(* Logix 5000 project; controller Joltek_RA_5069PLC002 vendor 1 type 14 code 226 rev 34.15; software revision 34.04 *) (continued)
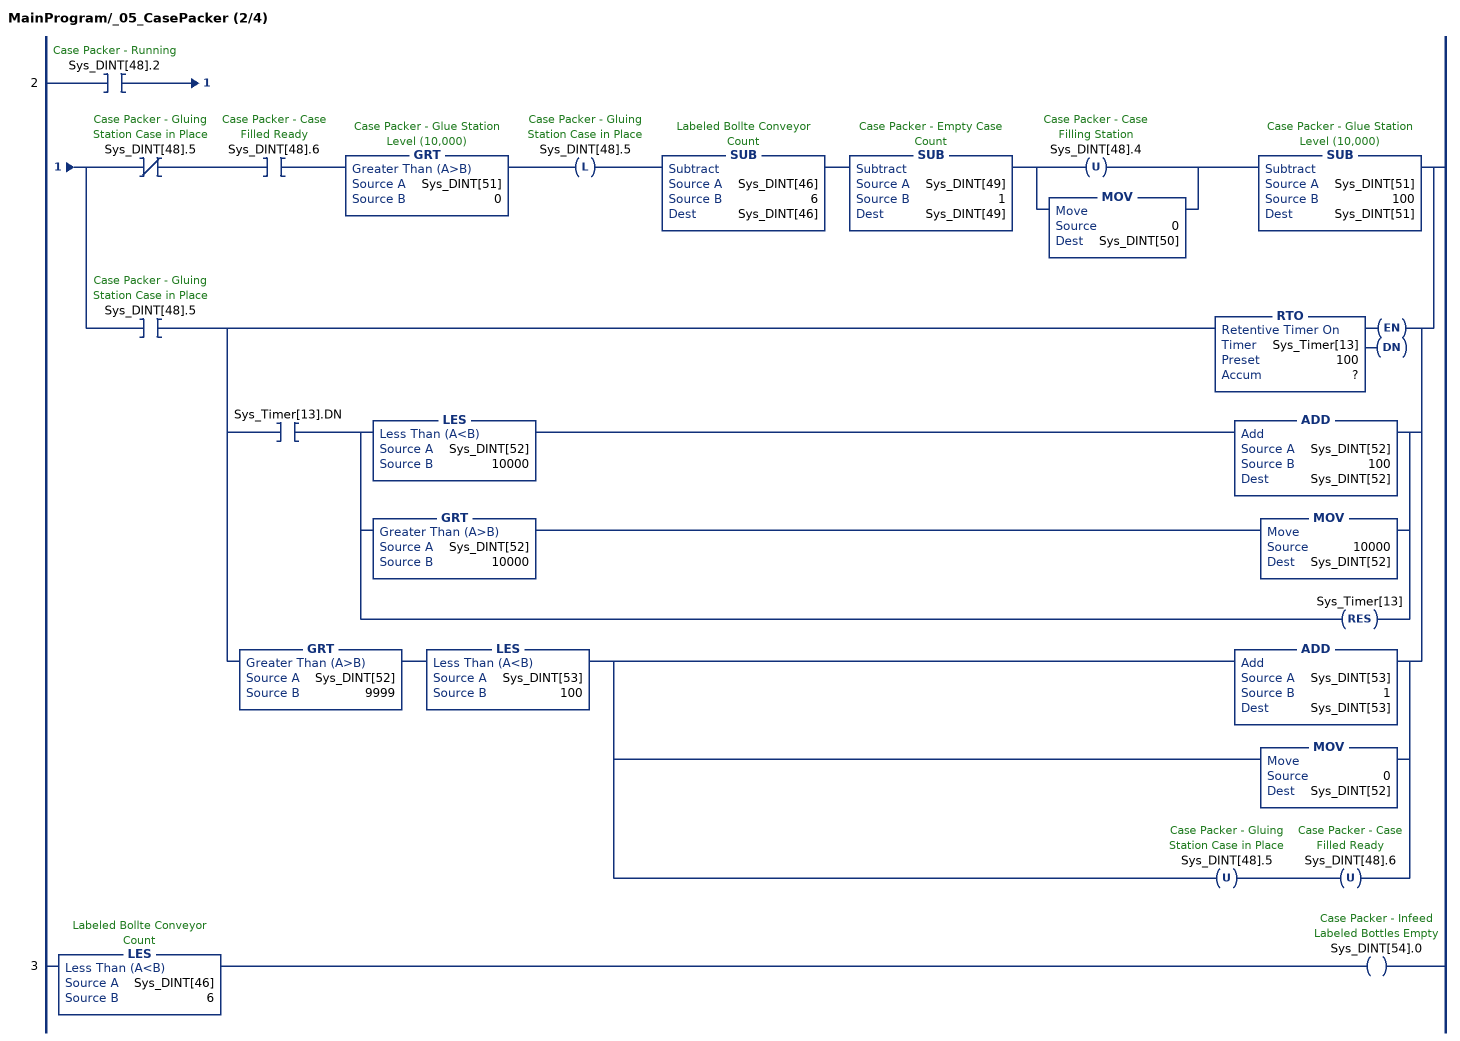
   2: XIC(Sys_DINT[48].2)[XIO(Sys_DINT[48].5) XIC(Sys_DINT[48].6) GRT(Sys_DINT[51],0) OTL(Sys_DINT[48].5) SUB(Sys_DINT[46],6,Sys_DINT[46]) SUB(Sys_DINT[49],1,Sys_DINT[49]) [OTU(Sys_DINT[48].4) ,MOV(0,Sys_DINT[50]) ] SUB(Sys_DINT[51],100,Sys_DINT[51]) ,XIC(Sys_DINT[48].5) [RTO(Sys_Timer[13],?,?) ,XIC(Sys_Timer[13].DN) [LES(Sys_DINT[52],10000) ADD(Sys_DINT[52],100,Sys_DINT[52]) ,GRT(Sys_DINT[52],10000) MOV(10000,Sys_DINT[52]) ,RES(Sys_Timer[13]) ] ,GRT(Sys_DINT[52],9999) LES(Sys_DINT[53],100) [ADD(Sys_DINT[53],1,Sys_DINT[53]) ,MOV(0,Sys_DINT[52]) ,OTU(Sys_DINT[48].5) OTU(Sys_DINT[48].6) ] ] ];
   3: LES(Sys_DINT[46],6)OTE(Sys_DINT[54].0);
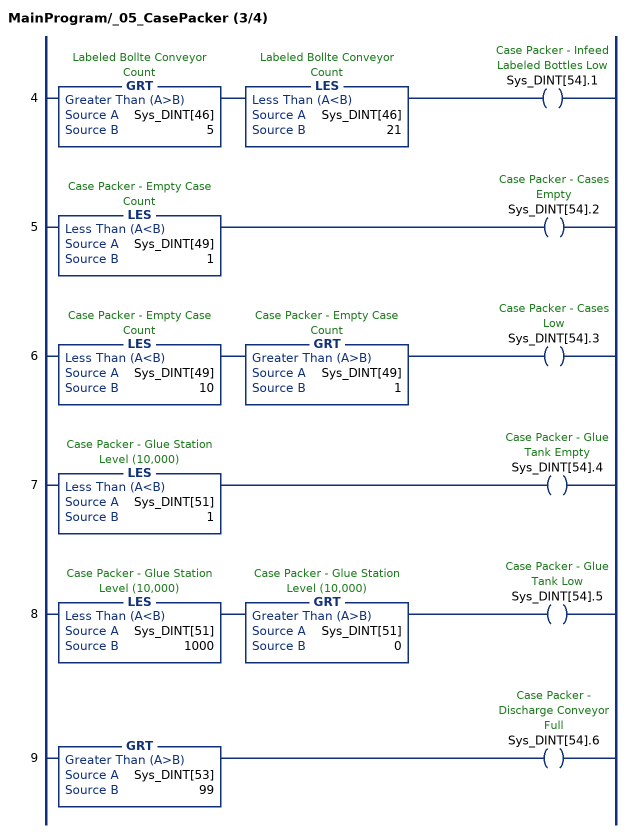
   4: GRT(Sys_DINT[46],5)LES(Sys_DINT[46],21)OTE(Sys_DINT[54].1);
   5: LES(Sys_DINT[49],1)OTE(Sys_DINT[54].2);
   6: LES(Sys_DINT[49],10)GRT(Sys_DINT[49],1)OTE(Sys_DINT[54].3);
   7: LES(Sys_DINT[51],1)OTE(Sys_DINT[54].4);
   8: LES(Sys_DINT[51],1000)GRT(Sys_DINT[51],0)OTE(Sys_DINT[54].5);
   9: GRT(Sys_DINT[53],99)OTE(Sys_DINT[54].6);
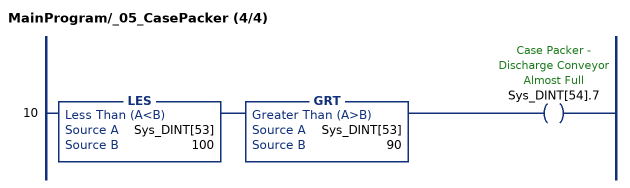
   10: LES(Sys_DINT[53],100)GRT(Sys_DINT[53],90)OTE(Sys_DINT[54].7);
END_ROUTINE

ROUTINE _06_Palletizer   (* ladder *)
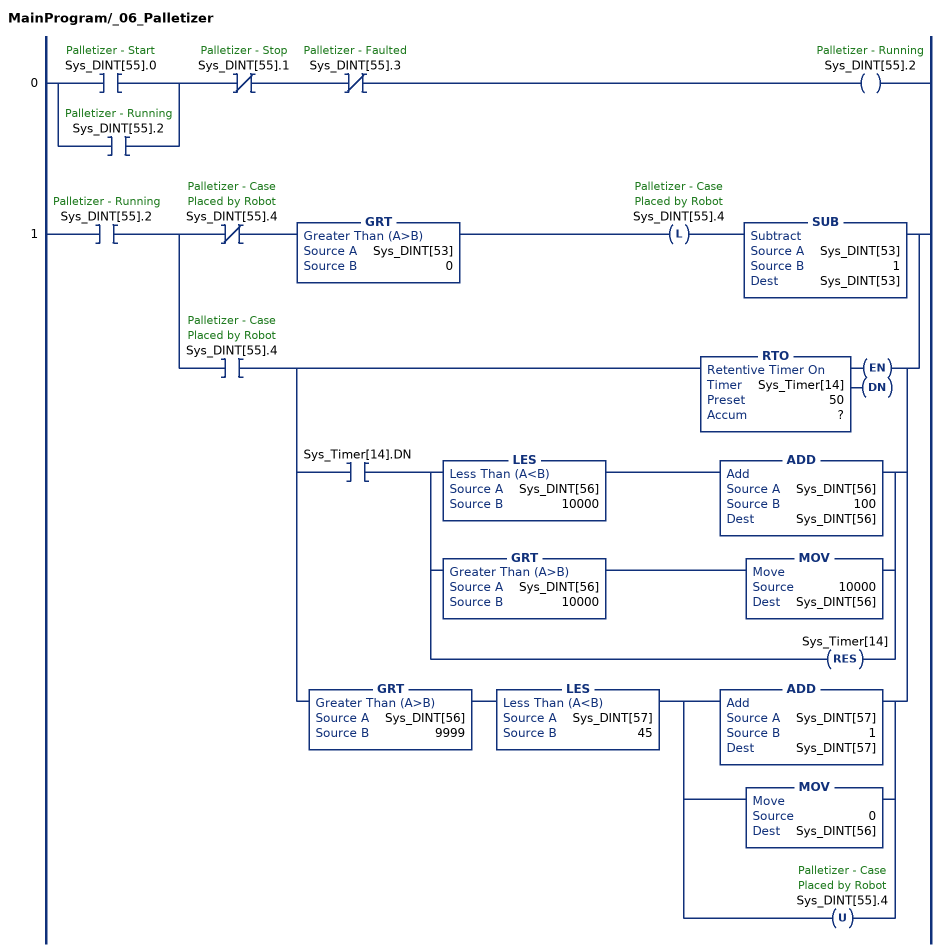
   0: [XIC(Sys_DINT[55].0) ,XIC(Sys_DINT[55].2) ]XIO(Sys_DINT[55].1)XIO(Sys_DINT[55].3)OTE(Sys_DINT[55].2);
   1: XIC(Sys_DINT[55].2)[XIO(Sys_DINT[55].4) GRT(Sys_DINT[53],0) OTL(Sys_DINT[55].4) SUB(Sys_DINT[53],1,Sys_DINT[53]) ,XIC(Sys_DINT[55].4) [RTO(Sys_Timer[14],?,?) ,XIC(Sys_Timer[14].DN) [LES(Sys_DINT[56],10000) ADD(Sys_DINT[56],100,Sys_DINT[56]) ,GRT(Sys_DINT[56],10000) MOV(10000,Sys_DINT[56]) ,RES(Sys_Timer[14]) ] ,GRT(Sys_DINT[56],9999) LES(Sys_DINT[57],45) [ADD(Sys_DINT[57],1,Sys_DINT[57]) ,MOV(0,Sys_DINT[56]) ,OTU(Sys_DINT[55].4) ] ] ];
END_ROUTINE

ROUTINE _50_HMI_Interface   (* ladder *)
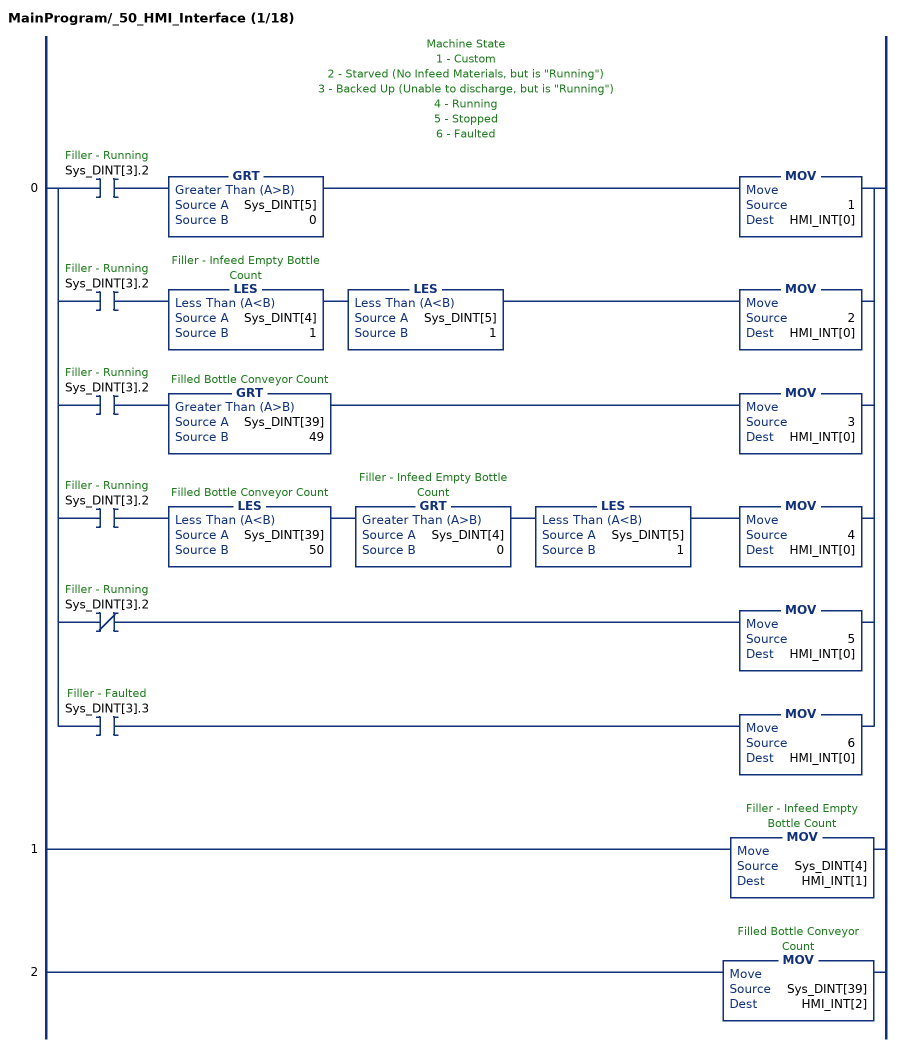
   // Machine State
   // 1 - Custom
   // 2 - Starved (No Infeed Materials, but is "Running")
   // 3 - Backed Up (Unable to discharge, but is "Running")
   // 4 - Running
   // 5 - Stopped
   // 6 - Faulted
   0: [XIC(Sys_DINT[3].2) GRT(Sys_DINT[5],0) MOV(1,HMI_INT[0]) ,XIC(Sys_DINT[3].2) LES(Sys_DINT[4],1) LES(Sys_DINT[5],1) MOV(2,HMI_INT[0]) ,XIC(Sys_DINT[3].2) GRT(Sys_DINT[39],49) MOV(3,HMI_INT[0]) ,XIC(Sys_DINT[3].2) LES(Sys_DINT[39],50) GRT(Sys_DINT[4],0) LES(Sys_DINT[5],1) MOV(4,HMI_INT[0]) ,XIO(Sys_DINT[3].2) MOV(5,HMI_INT[0]) ,XIC(Sys_DINT[3].3) MOV(6,HMI_INT[0]) ];
   1: MOV(Sys_DINT[4],HMI_INT[1]);
   2: MOV(Sys_DINT[39],HMI_INT[2]);
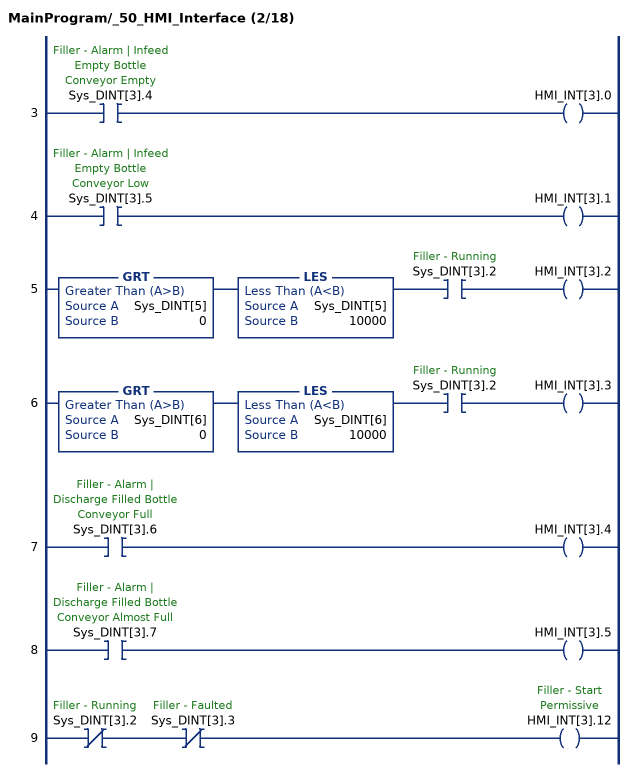
   3: XIC(Sys_DINT[3].4)OTE(HMI_INT[3].0);
   4: XIC(Sys_DINT[3].5)OTE(HMI_INT[3].1);
   5: GRT(Sys_DINT[5],0)LES(Sys_DINT[5],10000)XIC(Sys_DINT[3].2)OTE(HMI_INT[3].2);
   6: GRT(Sys_DINT[6],0)LES(Sys_DINT[6],10000)XIC(Sys_DINT[3].2)OTE(HMI_INT[3].3);
   7: XIC(Sys_DINT[3].6)OTE(HMI_INT[3].4);
   8: XIC(Sys_DINT[3].7)OTE(HMI_INT[3].5);
   9: XIO(Sys_DINT[3].2)XIO(Sys_DINT[3].3)OTE(HMI_INT[3].12);
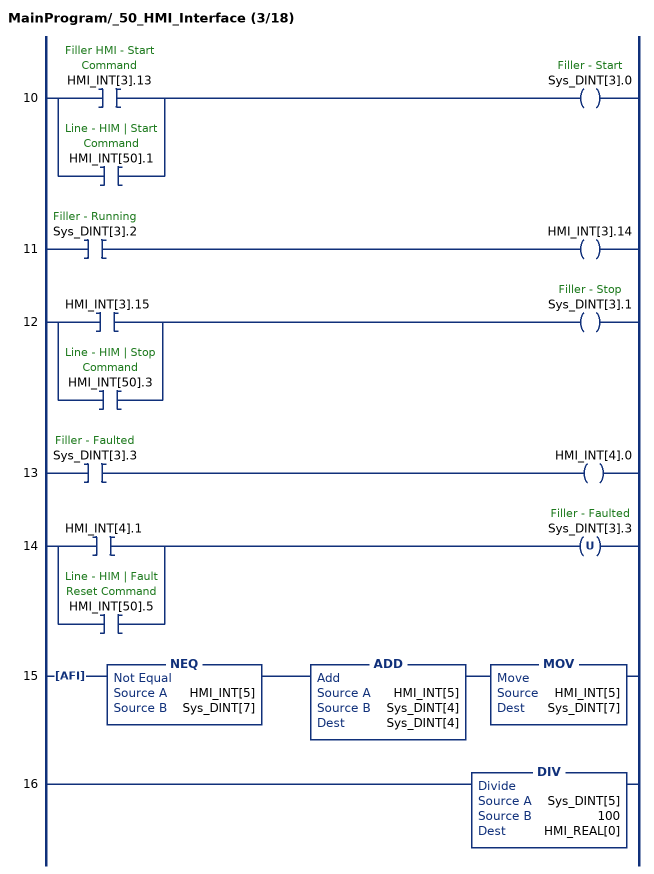
   10: [XIC(HMI_INT[3].13) ,XIC(HMI_INT[50].1) ]OTE(Sys_DINT[3].0);
   11: XIC(Sys_DINT[3].2)OTE(HMI_INT[3].14);
   12: [XIC(HMI_INT[3].15) ,XIC(HMI_INT[50].3) ]OTE(Sys_DINT[3].1);
   13: XIC(Sys_DINT[3].3)OTE(HMI_INT[4].0);
   14: [XIC(HMI_INT[4].1) ,XIC(HMI_INT[50].5) ]OTU(Sys_DINT[3].3);
   15: AFI()NEQ(HMI_INT[5],Sys_DINT[7])ADD(HMI_INT[5],Sys_DINT[4],Sys_DINT[4])MOV(HMI_INT[5],Sys_DINT[7]);
   16: DIV(Sys_DINT[5],100,HMI_REAL[0]);
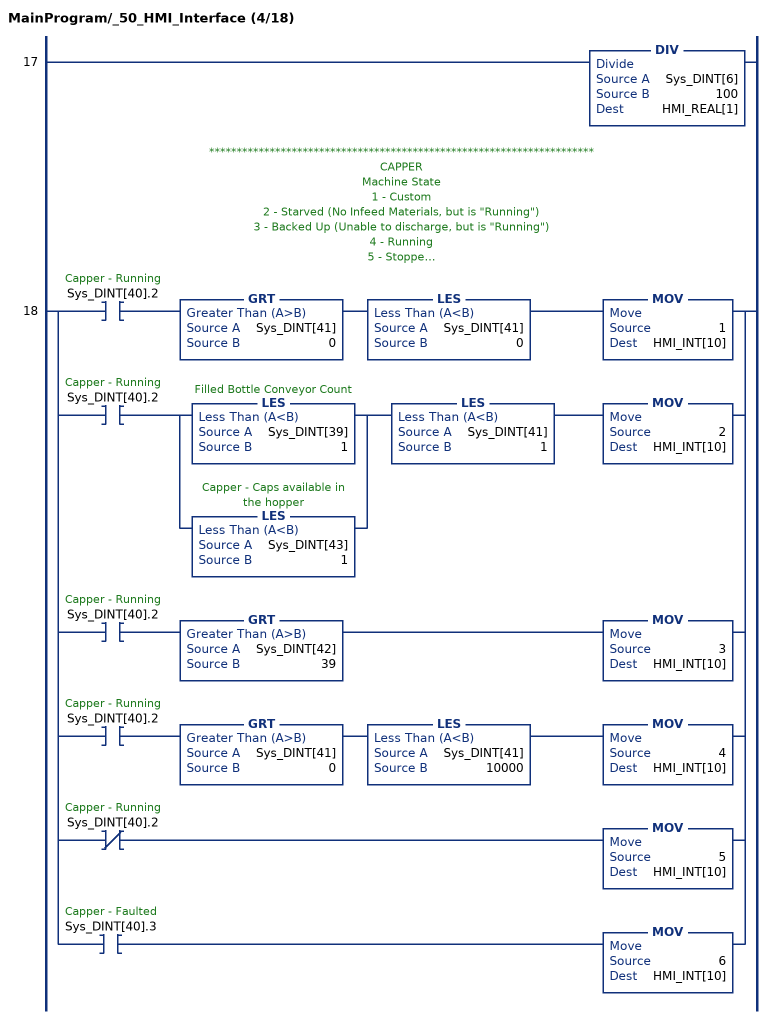
   17: DIV(Sys_DINT[6],100,HMI_REAL[1]);
   // **********************************************************************
   // CAPPER
   // Machine State
   // 1 - Custom
   // 2 - Starved (No Infeed Materials, but is "Running")
   // 3 - Backed Up (Unable to discharge, but is "Running")
   // 4 - Running
   // 5 - Stopped
   // 6 - Faulted
   18: [XIC(Sys_DINT[40].2) GRT(Sys_DINT[41],0) LES(Sys_DINT[41],0) MOV(1,HMI_INT[10]) ,XIC(Sys_DINT[40].2) [LES(Sys_DINT[39],1) ,LES(Sys_DINT[43],1) ] LES(Sys_DINT[41],1) MOV(2,HMI_INT[10]) ,XIC(Sys_DINT[40].2) GRT(Sys_DINT[42],39) MOV(3,HMI_INT[10]) ,XIC(Sys_DINT[40].2) GRT(Sys_DINT[41],0) LES(Sys_DINT[41],10000) MOV(4,HMI_INT[10]) ,XIO(Sys_DINT[40].2) MOV(5,HMI_INT[10]) ,XIC(Sys_DINT[40].3) MOV(6,HMI_INT[10]) ];
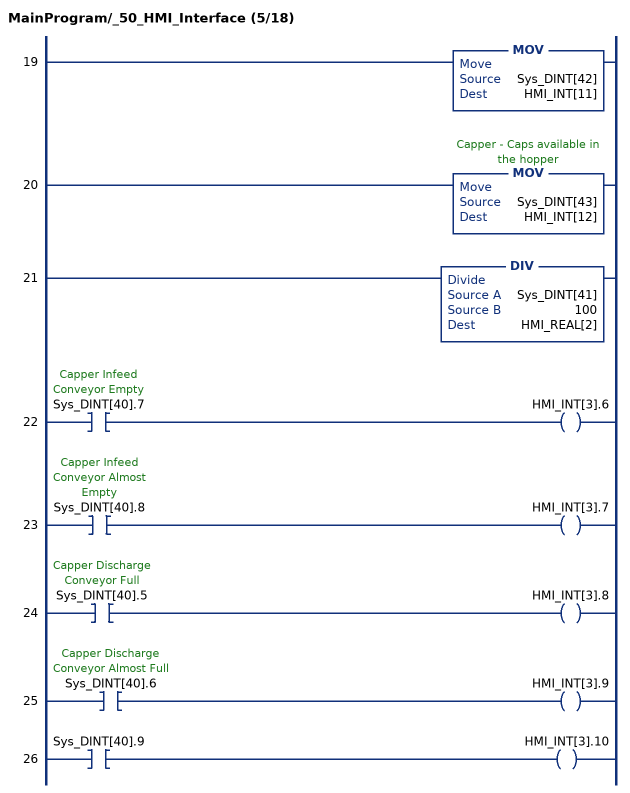
   19: MOV(Sys_DINT[42],HMI_INT[11]);
   20: MOV(Sys_DINT[43],HMI_INT[12]);
   21: DIV(Sys_DINT[41],100,HMI_REAL[2]);
   22: XIC(Sys_DINT[40].7)OTE(HMI_INT[3].6);
   23: XIC(Sys_DINT[40].8)OTE(HMI_INT[3].7);
   24: XIC(Sys_DINT[40].5)OTE(HMI_INT[3].8);
   25: XIC(Sys_DINT[40].6)OTE(HMI_INT[3].9);
   26: XIC(Sys_DINT[40].9)OTE(HMI_INT[3].10);
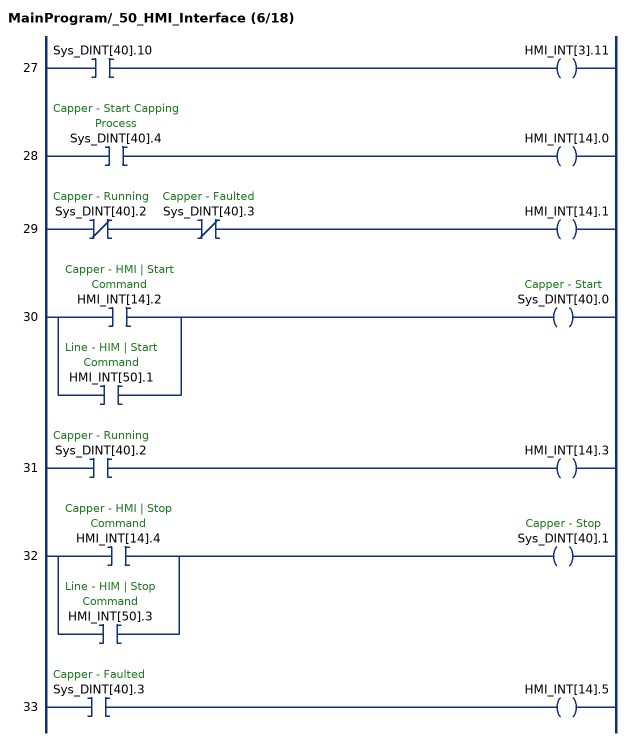
   27: XIC(Sys_DINT[40].10)OTE(HMI_INT[3].11);
   28: XIC(Sys_DINT[40].4)OTE(HMI_INT[14].0);
   29: XIO(Sys_DINT[40].2)XIO(Sys_DINT[40].3)OTE(HMI_INT[14].1);
   30: [XIC(HMI_INT[14].2) ,XIC(HMI_INT[50].1) ]OTE(Sys_DINT[40].0);
   31: XIC(Sys_DINT[40].2)OTE(HMI_INT[14].3);
   32: [XIC(HMI_INT[14].4) ,XIC(HMI_INT[50].3) ]OTE(Sys_DINT[40].1);
   33: XIC(Sys_DINT[40].3)OTE(HMI_INT[14].5);
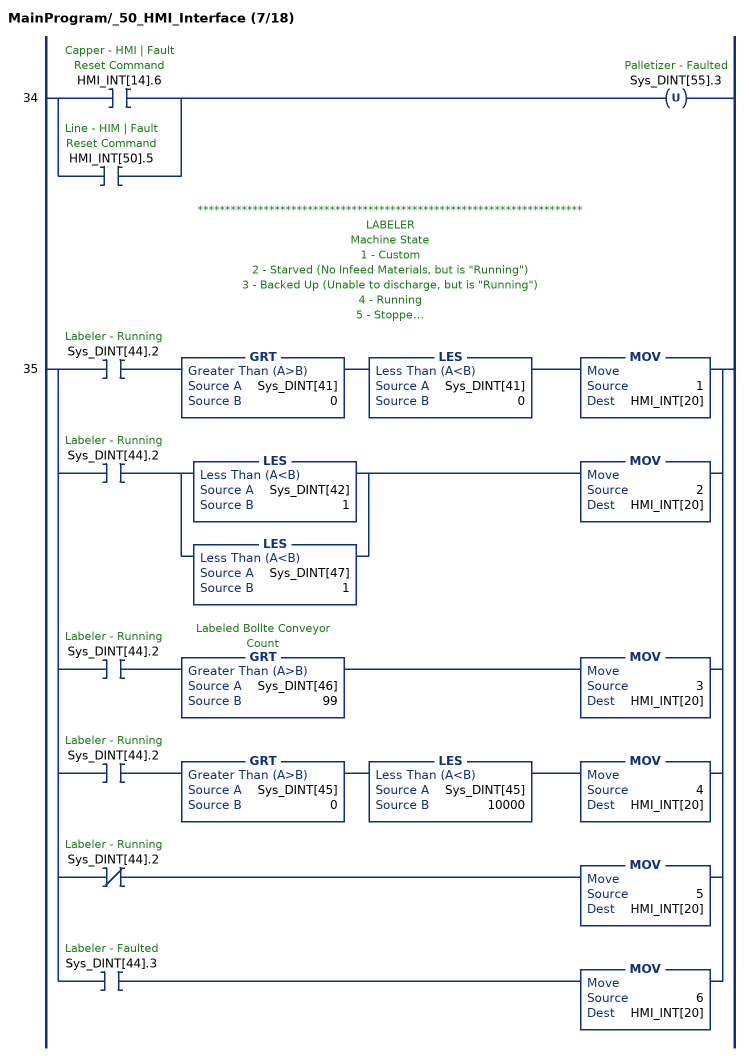
   34: [XIC(HMI_INT[14].6) ,XIC(HMI_INT[50].5) ]OTU(Sys_DINT[55].3);
   // **********************************************************************
   // LABELER
   // Machine State
   // 1 - Custom
   // 2 - Starved (No Infeed Materials, but is "Running")
   // 3 - Backed Up (Unable to discharge, but is "Running")
   // 4 - Running
   // 5 - Stopped
   // 6 - Faulted
   35: [XIC(Sys_DINT[44].2) GRT(Sys_DINT[41],0) LES(Sys_DINT[41],0) MOV(1,HMI_INT[20]) ,XIC(Sys_DINT[44].2) [LES(Sys_DINT[42],1) ,LES(Sys_DINT[47],1) ] MOV(2,HMI_INT[20]) ,XIC(Sys_DINT[44].2) GRT(Sys_DINT[46],99) MOV(3,HMI_INT[20]) ,XIC(Sys_DINT[44].2) GRT(Sys_DINT[45],0) LES(Sys_DINT[45],10000) MOV(4,HMI_INT[20]) ,XIO(Sys_DINT[44].2) MOV(5,HMI_INT[20]) ,XIC(Sys_DINT[44].3) MOV(6,HMI_INT[20]) ];
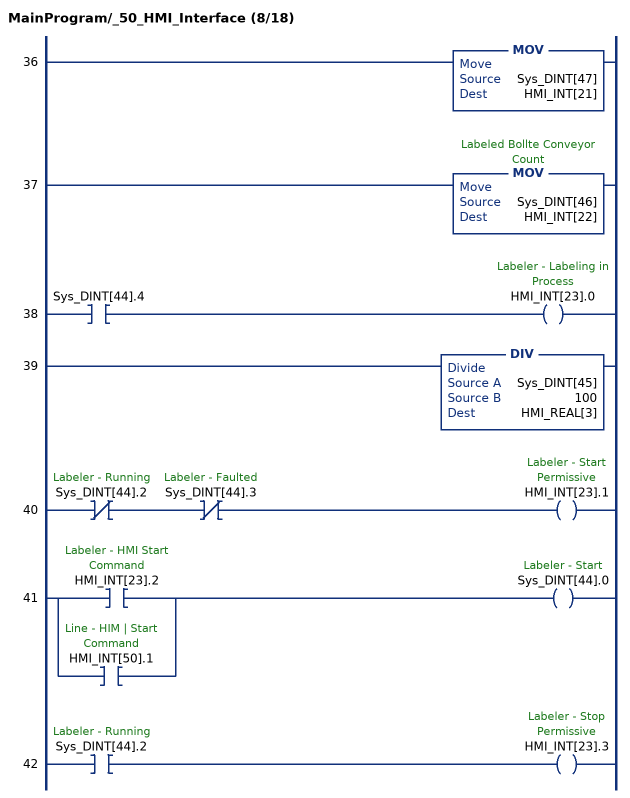
   36: MOV(Sys_DINT[47],HMI_INT[21]);
   37: MOV(Sys_DINT[46],HMI_INT[22]);
   38: XIC(Sys_DINT[44].4)OTE(HMI_INT[23].0);
   39: DIV(Sys_DINT[45],100,HMI_REAL[3]);
   40: XIO(Sys_DINT[44].2)XIO(Sys_DINT[44].3)OTE(HMI_INT[23].1);
   41: [XIC(HMI_INT[23].2) ,XIC(HMI_INT[50].1) ]OTE(Sys_DINT[44].0);
   42: XIC(Sys_DINT[44].2)OTE(HMI_INT[23].3);
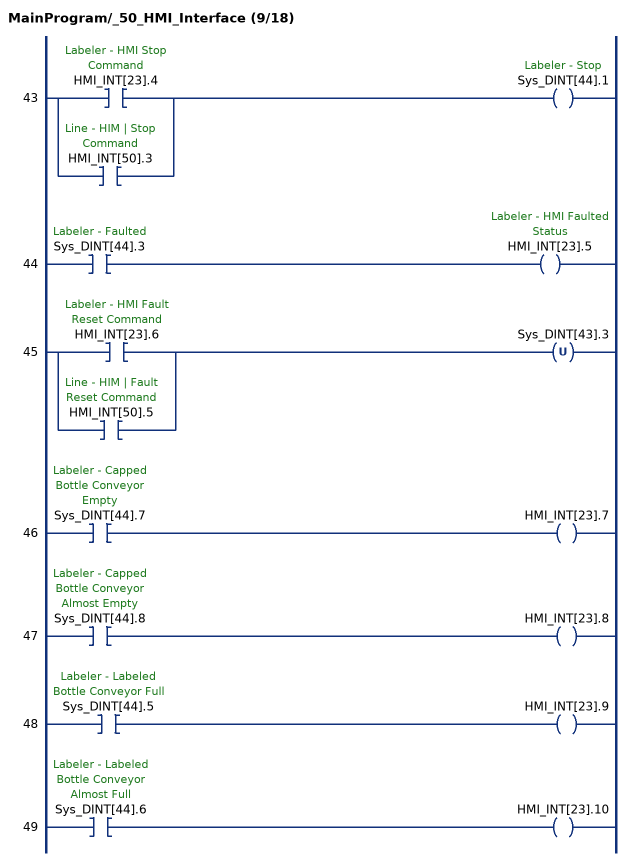
   43: [XIC(HMI_INT[23].4) ,XIC(HMI_INT[50].3) ]OTE(Sys_DINT[44].1);
   44: XIC(Sys_DINT[44].3)OTE(HMI_INT[23].5);
   45: [XIC(HMI_INT[23].6) ,XIC(HMI_INT[50].5) ]OTU(Sys_DINT[43].3);
   46: XIC(Sys_DINT[44].7)OTE(HMI_INT[23].7);
   47: XIC(Sys_DINT[44].8)OTE(HMI_INT[23].8);
   48: XIC(Sys_DINT[44].5)OTE(HMI_INT[23].9);
   49: XIC(Sys_DINT[44].6)OTE(HMI_INT[23].10);
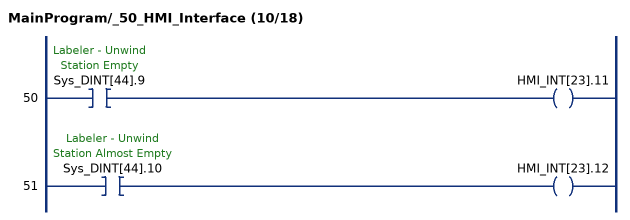
   50: XIC(Sys_DINT[44].9)OTE(HMI_INT[23].11);
   51: XIC(Sys_DINT[44].10)OTE(HMI_INT[23].12);
